(* Logix 5000 project; controller FV vendor 1 type 14 code 217 rev 31.11; software revision 31.00; part 55 of 63 *)
(* tags used below, declared in another part *)
   CWD : CHECKWORD_FLAGS;
   FV_B82 : INT[255];   // YSTFILL FL YST filling process flags
   FV_B86 : INT[255];   // YSTCIP FL YST CIP process flag s
   FV_B86_0_2_OutputBit : BOOL;
   FV_N144 : INT[255];   // YST1 DATA
   FV_N145 : INT[255];   // YST2 DATA
   FV_N80 : INT[255];   // YSTFILL<PC YST filling data fro m PC
   FV_N81 : INT[255];   // YSTFILL>PC YST filling process data to PC and contr ol regs.
   FV_N84 : INT[255];   // YSTCIP<PC YST CIP data from PC
   FV_N85 : INT[255];   // YSTCIP>PC YST CIP process data to PC and control r egs.
   FV_N88 : INT[255];   // YSP COMMS Data transferred to/ from yeast press PLC
   FV_R2V1 : PlantItem;   // R2V1
   FV_R2V2 : PlantItem;   // R2V2
   FV_T83 : TIMER[5];
   FV_T87 : TIMER[2];
   FV_T89 : TIMER[5];
   FV_WYTR1 : PlantItem;   // WYTR1
   FV_WYTR2 : PlantItem;   // WYTR2
   FV_Yeast_Press_Blunger_Comms : MESSAGE;
   FV_YST1_HL_SP : DINT;
   FV_YST2_HL_SP : DINT;
   MV_YST_Levels : REAL[2];
   YST_BL_PMP_ON : BOOL;   // Blunger Pump
   YST_CIP_Conns_Confirmed : BOOL;
   YST_Confirm_CIP_connected : BOOL;
(* FV_Common, continued *)

ROUTINE FV_YSP_COMMS_88   (* ladder *)
   // Communications with Yeast Press PLC routine
   0: XIO(FV_T89[0].DN)TON(FV_T89[0],?,?);
   1: XIC(FV_T89[0].DN)MSG(FV_Yeast_Press_Blunger_Comms);
   2: XIO(FV_N88[10].0)[OTE(FV_N88[0].0) ,TON(FV_T89[1],?,?) ];
   3: XIC(FV_N88[10].0)TON(FV_T89[2],?,?);
   4: [XIC(FV_T89[1].DN) ,XIC(FV_T89[2].DN) ]OTE(FV_N88[20].0);
END_ROUTINE

ROUTINE FV_YSTCIP_CP_85   (* ladder *)
   // YST CIP Command Processor Reset current step on first scan
   0: XIC(S:FS)CLR(FV_N85[16]);
   // Step 0: reset
   1: EQU(FV_N85[16],0)MCR();
   2: [OTU(FV_B86[0].0) ,OTU(FV_B86[0].1) ];
   3: [FLL(0,FV_N85[0],16) ,FLL(-32768,FV_N84[1],7) ,CLR(FV_N84[0]) ];
   4: MOV(1,FV_N85[16]);
   5: MCR();
   // Step 1: wait for start from PC
   6: EQU(FV_N85[16],1)MCR();
   7: MOV(1,FV_N85[0]);
   // Allow startup if any YST is inactive or on storage
   8: [[EQU(FV_N144[0],0) ,EQU(FV_N144[0],5) ] NEQ(FV_N145[0],1) ,[EQU(FV_N145[0],0) ,EQU(FV_N145[0],5) ] NEQ(FV_N144[0],1) ]OTE(FV_N85[2].0);
   9: XIC(FV_N85[2].0)XIC(FV_N84[0].0)MOV(2,FV_N85[16]);
   10: MCR();
   // Step 2: startup in progress
   11: EQU(FV_N85[16],2)MCR();
   // If YST1 selected and no other YST1 startup in progress enable CIP start flag
   12: EQU(FV_N84[1],1)[EQU(FV_N144[0],0) ,EQU(FV_N144[0],5) ][EQU(FV_N144[4],0) ,XIC(FV_N144[4].3) ]OTE(FV_N144[4].3);
   13: EQU(FV_N84[1],2)[EQU(FV_N145[0],0) ,EQU(FV_N145[0],5) ][EQU(FV_N145[4],0) ,XIC(FV_N145[4].3) ]OTE(FV_N145[4].3);
   14: [XIC(FV_N144[4].3) ,XIC(FV_N145[4].3) ]OTE(FV_N85[2].1);
   15: TON(FV_T87[0],?,?);
   16: [XIC(FV_N84[0].15) ,XIC(FV_T87[0].DN) ]CLR(FV_N85[16]);
   17: XIC(FV_N84[0].1)XIC(FV_N85[2].1)[MOV(3,FV_N85[16]) ,CLR(FV_N84[0]) ];
   18: MCR();
   // Step 3: complete startup
   19: EQU(FV_N85[16],3)MCR();
   // If selected YST is YST1 set YST1's status to CIP
   20: EQU(FV_N84[1],1)MOV(3,FV_N144[0]);
   // If selected YST is YST2 set YST2's status tto CIP
   21: EQU(FV_N84[1],2)MOV(3,FV_N145[0]);
   // Activate YST CIP process
   22: [MOV(2,FV_N85[0]) ,OTL(FV_B86[0].0) ,OTL(FV_B86[0].1) ,OTL(FV_N85[2].2) ,MOV(10,FV_N85[1]) ,MOV(10,FV_N85[3]) ];
   23: [MOV(-1,FV_N85[16]) ,CLR(FV_N84[0]) ];
   24: MCR();
   // YST CIP stop button
   25: XIC(FV_N85[2].2)XIC(FV_N84[0].2)MCR();
   26: [OTU(FV_B86[0].1) ,OTU(FV_N85[2].2) ,OTL(FV_N85[2].3) ,OTL(FV_N85[2].4) ];
   27: [MOV(3,FV_N85[0]) ,MOV(0,FV_N85[1]) ,CLR(FV_N84[0]) ];
   28: MCR();
   // YST CIP continue button
   29: XIC(FV_N85[2].3)XIC(FV_N84[0].3)MCR();
   30: [OTL(FV_B86[0].1) ,OTL(FV_N85[2].2) ,OTU(FV_N85[2].3) ,OTU(FV_N85[2].4) ];
   31: [FLL(0,FV_N85[4],4) ,MOV(2,FV_N85[0]) ,MOV(FV_N85[3],FV_N85[1]) ,CLR(FV_N84[0]) ];
   32: MCR();
   // YST CIP abort button
   33: XIC(FV_N85[2].4)XIC(FV_N84[0].4)MCR();
   34: OTU(FV_B86[0].0);
   // Set current YST's operation to none
   35: JSR(FV_Set_FV_Datafile_Value,3,0,FV_N85[15],0);
   36: [CLR(FV_N85[16]) ,CLR(FV_N84[0]) ];
   37: MCR();
   // Copy current step to PC display register
   38: XIC(FV_B86[0].1)MOV(FV_N85[1],FV_N85[9]);
END_ROUTINE

ROUTINE FV_YSTCIP_MC_84   (* ladder *)
   // YST CIP master control program YST CIP command processor
   0: JSR(FV_YSTCIP_CP_85,0);
   // YST CIP process control program
   1: XIC(FV_B86[0].0)JSR(FV_YSTCIP_PR_86,0);
   // Postscan YST CIP program
   2: XIO(FV_B86[0].0)OSR(FV_B86[0].2,FV_B86_0_2_OutputBit)XIC(FV_B86_0_2_OutputBit)JSR(FV_YSTCIP_PR_86,0);
   // Keep CIP valve open to prevent buildup of pressure in YST1
   3: XIO(FV_B86[0].1)[EQU(FV_N144[0],5) ,XIC(FV_N81[2].3) EQU(FV_N144[0],1) ]OTE(FV_R2V1.DriveBits.2);
   // Keep CIP valve open to prevent buildup of pressure in YST2
   4: XIO(FV_B86[0].1)[EQU(FV_N145[0],5) ,XIC(FV_N81[2].3) EQU(FV_N145[0],1) ]OTE(FV_R2V2.DriveBits.2);
END_ROUTINE

ROUTINE FV_YSTCIP_PR_86   (* ladder *)
   // YST Filling Process Control Program Step 10: Initialise
   0: XIC(FV_B86[0].1)EQU(FV_N85[1],10)MCR();
   1: [OTE(YST_Confirm_CIP_connected) ,XIC(YST_CIP_Conns_Confirmed) MOV(11,FV_N85[1]) ];
   2: MCR();
   // YST CIP Process Control Program Step 10: Initialise
   3: XIC(FV_B86[0].1)EQU(FV_N85[1],11)MCR();
   4: MOV(10,FV_N85[3]);
   // Initialise pointer to current YST's data and attemperation files
   5: [ADD(FV_N84[1],143,FV_N85[15]) ,ADD(FV_N84[1],138,FV_N85[14]) ];
   // Set rouser mode to automatic
   6: JSR(FV_Set_FV_Datafile_Value,3,0,FV_N85[15],3);
   // Stop attemperation control on selected YST
   7: [JSR(FV_Set_FV_Datafile_Value,3,0,FV_N85[14],24) ,JSR(FV_Set_FV_Datafile_Value,3,0,FV_N85[14],26) JSR(FV_Set_FV_Datafile_Value,3,0,FV_N85[14],27) JSR(FV_Set_FV_Datafile_Value,3,0,FV_N85[14],28) JSR(FV_Set_FV_Datafile_Value,3,0,FV_N85[14],29) JSR(FV_Set_FV_Datafile_Value,3,0,FV_N85[14],30) JSR(FV_Set_FV_Datafile_Value,3,0,FV_N85[14],31) ];
   8: MOV(20,FV_N85[1]);
   9: MCR();
   // Step 20: Open CIP route
   10: EQU(FV_N85[1],20)MCR();
   11: MOV(20,FV_N85[3]);
   12: [EQU(FV_N84[1],1) OTE(FV_R2V1.DriveBits.0) ,EQU(FV_N84[1],2) OTE(FV_R2V2.DriveBits.0) ];
   13: [OTE(FV_N85[2].5) ,XIC(FV_N84[0].5) MOV(30,FV_N85[1]) ];
   14: MCR();
   // Step 30: reset YST
   15: EQU(FV_N85[1],30)MCR();
   // Unlatch current YST dirty flag
   16: JSR(FV_Clear_Flag_In_FV_Datafile,3,FV_N85[15],1,0);
   17: [JSR(FV_Set_FV_Datafile_Value,3,0,FV_N85[15],0) ,CLR(FV_N85[16]) ];
   18: MCR();
   // Check for alarms while running
   19: XIC(FV_B86[0].1)MCR();
   20: [EQU(FV_N84[1],1) [XIC(FV_R2V1.CW.[CWD.FAULT]) ,XIC(FV_WYTR1.CW.[CWD.FAULT]) ] ,EQU(FV_N84[1],2) [XIC(FV_R2V2.CW.[CWD.FAULT]) ,XIC(FV_WYTR2.CW.[CWD.FAULT]) ] ,GRT(FV_N85[4],0) ]OTU(FV_B86[0].1);
   21: XIO(FV_B86[0].1)[MOV(4,FV_N85[0]) ,OTU(FV_N85[2].2) ,OTL(FV_N85[2].3) ,OTL(FV_N85[2].4) ,MOV(0,FV_N85[1]) ];
   22: MCR();
END_ROUTINE

ROUTINE FV_YSTFILL_CP_81   (* ladder *)
   // YST Filling Command Processor Reset current step on first scan
   0: XIC(S:FS)CLR(FV_N81[16]);
   // Step 0: reset
   1: EQU(FV_N81[16],0)MCR();
   2: [OTU(FV_B82[0].0) ,OTU(FV_B82[0].1) ];
   3: [FLL(0,FV_N81[0],16) ,FLL(-32768,FV_N80[1],7) ,CLR(FV_N80[0]) ];
   4: MOV(1,FV_N81[16]);
   5: MCR();
   // Step 1: wait for start from PC
   6: EQU(FV_N81[16],1)MCR();
   7: MOV(1,FV_N81[0]);
   // Allow startup if any YST is inactive or on storage
   8: [[EQU(FV_N144[0],0) ,EQU(FV_N144[0],5) ] NEQ(FV_N145[0],3) LEQ(MV_YST_Levels[0],FV_YST1_HL_SP) ,[EQU(FV_N145[0],0) ,EQU(FV_N145[0],5) ] NEQ(FV_N144[0],3) LEQ(MV_YST_Levels[1],FV_YST2_HL_SP) ]OTE(FV_N81[2].0);
   9: XIC(FV_N81[2].0)XIC(FV_N80[0].0)MOV(2,FV_N81[16]);
   10: MCR();
   // Step 2: startup in progress
   11: EQU(FV_N81[16],2)MCR();
   // If YST1 selected and no other YST1 startup in progress enable filling start flag
   12: EQU(FV_N80[1],1)[EQU(FV_N144[0],0) ,EQU(FV_N144[0],5) ][EQU(FV_N144[4],0) ,XIC(FV_N144[4].1) ]OTE(FV_N144[4].1);
   // If YST2 selected and no other YST2 startup in progress enable filling start flag
   13: EQU(FV_N80[1],2)[EQU(FV_N145[0],0) ,EQU(FV_N145[0],5) ][EQU(FV_N145[4],0) ,XIC(FV_N145[4].1) ]OTE(FV_N145[4].1);
   // Enable start button of selected YST could be locked
   14: [XIC(FV_N144[4].1) ,XIC(FV_N145[4].1) ]OTE(FV_N81[2].1);
   15: TON(FV_T83[0],?,?);
   16: [XIC(FV_N80[0].15) ,XIC(FV_T83[0].DN) ]CLR(FV_N81[16]);
   17: XIC(FV_N80[0].1)XIC(FV_N81[2].1)[MOV(3,FV_N81[16]) ,CLR(FV_N80[0]) ];
   18: MCR();
   // Step 3: complete startup
   19: EQU(FV_N81[16],3)MCR();
   // Set appropriate YST's status to filling
   20: EQU(FV_N80[1],1)MOV(1,FV_N144[0]);
   21: EQU(FV_N80[1],2)MOV(1,FV_N145[0]);
   // Activate YST filling process
   22: [MOV(2,FV_N81[0]) ,OTL(FV_B82[0].0) ,OTL(FV_B82[0].1) ,OTL(FV_N81[2].2) ,MOV(10,FV_N81[1]) ,MOV(10,FV_N81[3]) ];
   23: [MOV(-1,FV_N81[16]) ,CLR(FV_N80[0]) ];
   24: MCR();
   // YST filling stop button
   25: XIC(FV_N81[2].2)XIC(FV_N80[0].2)MCR();
   26: [OTU(FV_B82[0].1) ,OTU(FV_N81[2].2) ,OTL(FV_N81[2].3) ,OTL(FV_N81[2].4) ,OTU(YST_BL_PMP_ON) ];
   27: [MOV(3,FV_N81[0]) ,MOV(0,FV_N81[1]) ,CLR(FV_N80[0]) ];
   28: MCR();
   // YST filling continue button
   29: XIC(FV_N81[2].3)XIC(FV_N80[0].3)MCR();
   30: [OTL(FV_B82[0].1) ,OTL(FV_N81[2].2) ,OTU(FV_N81[2].3) ,OTU(FV_N81[2].4) ];
   31: [FLL(0,FV_N81[4],4) ,MOV(2,FV_N81[0]) ,MOV(FV_N81[3],FV_N81[1]) ,CLR(FV_N80[0]) ];
   32: MCR();
   // YST filling abort button
   33: XIC(FV_N81[2].4)XIC(FV_N80[0].4)MCR();
